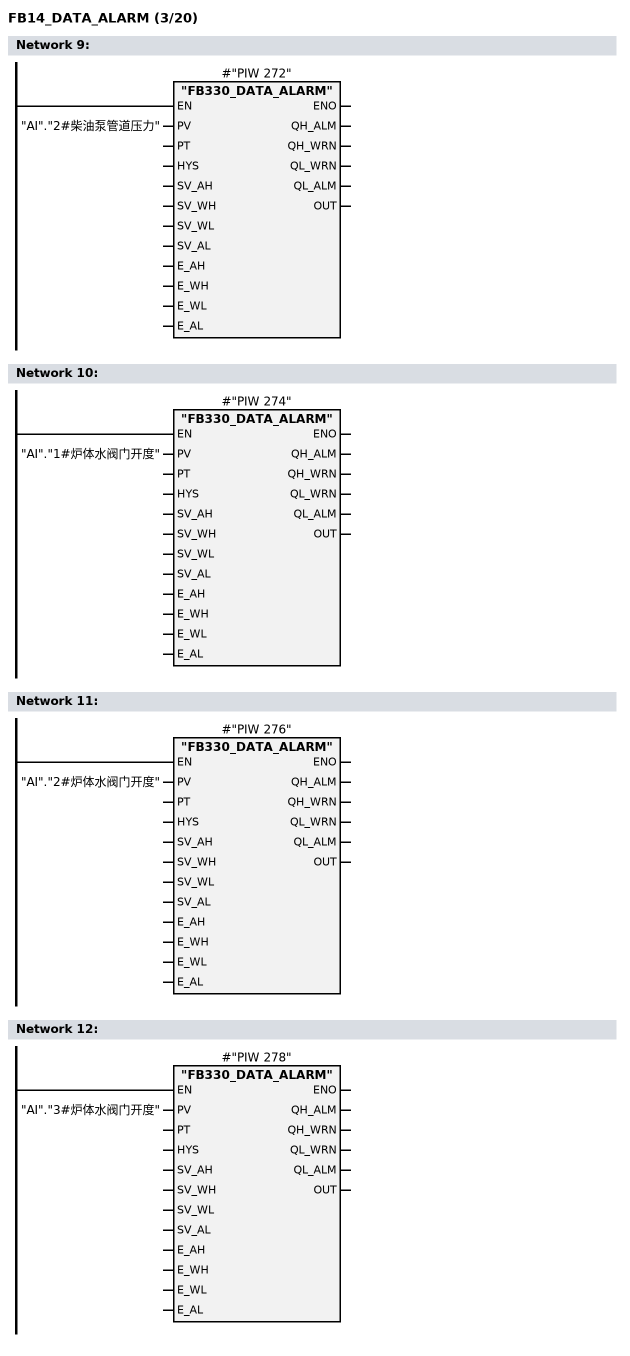
   RUNG wire#powerrail
      #"PIW 272"(PV := "AI"."2#柴油泵管道压力", PT :=, HYS :=, SV_AH :=, SV_WH :=, SV_WL :=, SV_AL :=, E_AH :=, E_WH :=, E_WL :=, E_AL :=, QH_ALM =>, QH_WRN =>, QL_WRN =>, QL_ALM =>, OUT =>)
   END_RUNG
   // the same network as SCL:
   #"PIW 272"(PV := "AI"."2#柴油泵管道压力");   // "FB330_DATA_ALARM"
END_REGION

REGION Network 10
   RUNG wire#powerrail
      #"PIW 274"(PV := "AI"."1#炉体水阀门开度", PT :=, HYS :=, SV_AH :=, SV_WH :=, SV_WL :=, SV_AL :=, E_AH :=, E_WH :=, E_WL :=, E_AL :=, QH_ALM =>, QH_WRN =>, QL_WRN =>, QL_ALM =>, OUT =>)
   END_RUNG
   // the same network as SCL:
   #"PIW 274"(PV := "AI"."1#炉体水阀门开度");   // "FB330_DATA_ALARM"
END_REGION

REGION Network 11
   RUNG wire#powerrail
      #"PIW 276"(PV := "AI"."2#炉体水阀门开度", PT :=, HYS :=, SV_AH :=, SV_WH :=, SV_WL :=, SV_AL :=, E_AH :=, E_WH :=, E_WL :=, E_AL :=, QH_ALM =>, QH_WRN =>, QL_WRN =>, QL_ALM =>, OUT =>)
   END_RUNG
   // the same network as SCL:
   #"PIW 276"(PV := "AI"."2#炉体水阀门开度");   // "FB330_DATA_ALARM"
END_REGION

REGION Network 12
   RUNG wire#powerrail
      #"PIW 278"(PV := "AI"."3#炉体水阀门开度", PT :=, HYS :=, SV_AH :=, SV_WH :=, SV_WL :=, SV_AL :=, E_AH :=, E_WH :=, E_WL :=, E_AL :=, QH_ALM =>, QH_WRN =>, QL_WRN =>, QL_ALM =>, OUT =>)
   END_RUNG
   // the same network as SCL:
   #"PIW 278"(PV := "AI"."3#炉体水阀门开度");   // "FB330_DATA_ALARM"
END_REGION

REGION Network 13
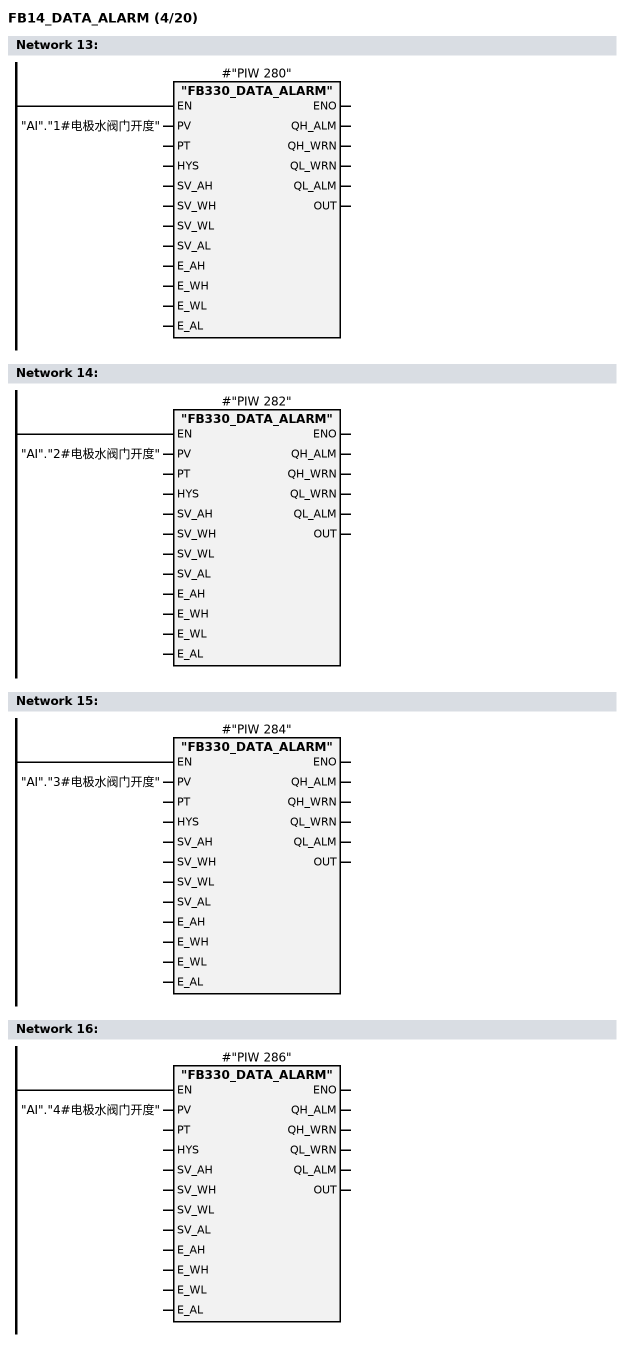
   RUNG wire#powerrail
      #"PIW 280"(PV := "AI"."1#电极水阀门开度", PT :=, HYS :=, SV_AH :=, SV_WH :=, SV_WL :=, SV_AL :=, E_AH :=, E_WH :=, E_WL :=, E_AL :=, QH_ALM =>, QH_WRN =>, QL_WRN =>, QL_ALM =>, OUT =>)
   END_RUNG
   // the same network as SCL:
   #"PIW 280"(PV := "AI"."1#电极水阀门开度");   // "FB330_DATA_ALARM"
END_REGION

REGION Network 14
   RUNG wire#powerrail
      #"PIW 282"(PV := "AI"."2#电极水阀门开度", PT :=, HYS :=, SV_AH :=, SV_WH :=, SV_WL :=, SV_AL :=, E_AH :=, E_WH :=, E_WL :=, E_AL :=, QH_ALM =>, QH_WRN =>, QL_WRN =>, QL_ALM =>, OUT =>)
   END_RUNG
   // the same network as SCL:
   #"PIW 282"(PV := "AI"."2#电极水阀门开度");   // "FB330_DATA_ALARM"
END_REGION

REGION Network 15
   RUNG wire#powerrail
      #"PIW 284"(PV := "AI"."3#电极水阀门开度", PT :=, HYS :=, SV_AH :=, SV_WH :=, SV_WL :=, SV_AL :=, E_AH :=, E_WH :=, E_WL :=, E_AL :=, QH_ALM =>, QH_WRN =>, QL_WRN =>, QL_ALM =>, OUT =>)
   END_RUNG
   // the same network as SCL:
   #"PIW 284"(PV := "AI"."3#电极水阀门开度");   // "FB330_DATA_ALARM"
END_REGION

REGION Network 16
   RUNG wire#powerrail
      #"PIW 286"(PV := "AI"."4#电极水阀门开度", PT :=, HYS :=, SV_AH :=, SV_WH :=, SV_WL :=, SV_AL :=, E_AH :=, E_WH :=, E_WL :=, E_AL :=, QH_ALM =>, QH_WRN =>, QL_WRN =>, QL_ALM =>, OUT =>)
   END_RUNG
   // the same network as SCL:
   #"PIW 286"(PV := "AI"."4#电极水阀门开度");   // "FB330_DATA_ALARM"
END_REGION

REGION Network 17
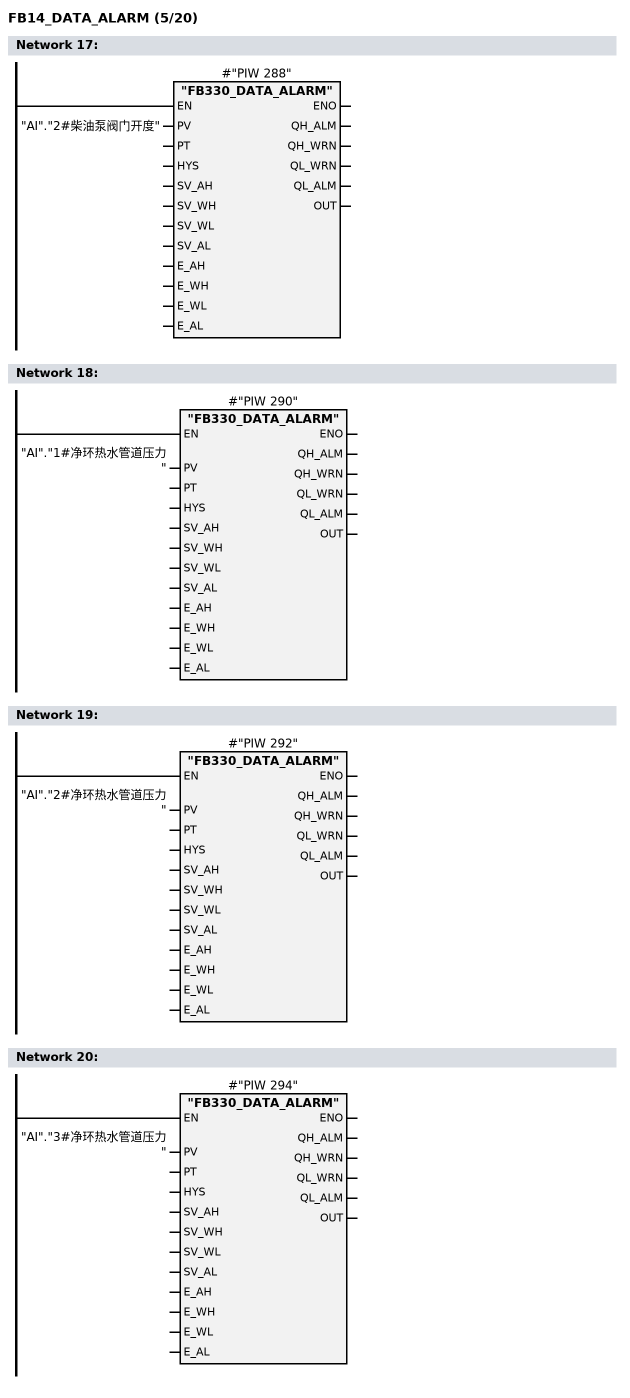
   RUNG wire#powerrail
      #"PIW 288"(PV := "AI"."2#柴油泵阀门开度", PT :=, HYS :=, SV_AH :=, SV_WH :=, SV_WL :=, SV_AL :=, E_AH :=, E_WH :=, E_WL :=, E_AL :=, QH_ALM =>, QH_WRN =>, QL_WRN =>, QL_ALM =>, OUT =>)
   END_RUNG
   // the same network as SCL:
   #"PIW 288"(PV := "AI"."2#柴油泵阀门开度");   // "FB330_DATA_ALARM"
END_REGION

REGION Network 18
   RUNG wire#powerrail
      #"PIW 290"(PV := "AI"."1#净环热水管道压力", PT :=, HYS :=, SV_AH :=, SV_WH :=, SV_WL :=, SV_AL :=, E_AH :=, E_WH :=, E_WL :=, E_AL :=, QH_ALM =>, QH_WRN =>, QL_WRN =>, QL_ALM =>, OUT =>)
   END_RUNG
   // the same network as SCL:
   #"PIW 290"(PV := "AI"."1#净环热水管道压力");   // "FB330_DATA_ALARM"
END_REGION

REGION Network 19
   RUNG wire#powerrail
      #"PIW 292"(PV := "AI"."2#净环热水管道压力", PT :=, HYS :=, SV_AH :=, SV_WH :=, SV_WL :=, SV_AL :=, E_AH :=, E_WH :=, E_WL :=, E_AL :=, QH_ALM =>, QH_WRN =>, QL_WRN =>, QL_ALM =>, OUT =>)
   END_RUNG
   // the same network as SCL:
   #"PIW 292"(PV := "AI"."2#净环热水管道压力");   // "FB330_DATA_ALARM"
END_REGION

REGION Network 20
   RUNG wire#powerrail
      #"PIW 294"(PV := "AI"."3#净环热水管道压力", PT :=, HYS :=, SV_AH :=, SV_WH :=, SV_WL :=, SV_AL :=, E_AH :=, E_WH :=, E_WL :=, E_AL :=, QH_ALM =>, QH_WRN =>, QL_WRN =>, QL_ALM =>, OUT =>)
   END_RUNG
   // the same network as SCL:
   #"PIW 294"(PV := "AI"."3#净环热水管道压力");   // "FB330_DATA_ALARM"
END_REGION

REGION Network 21
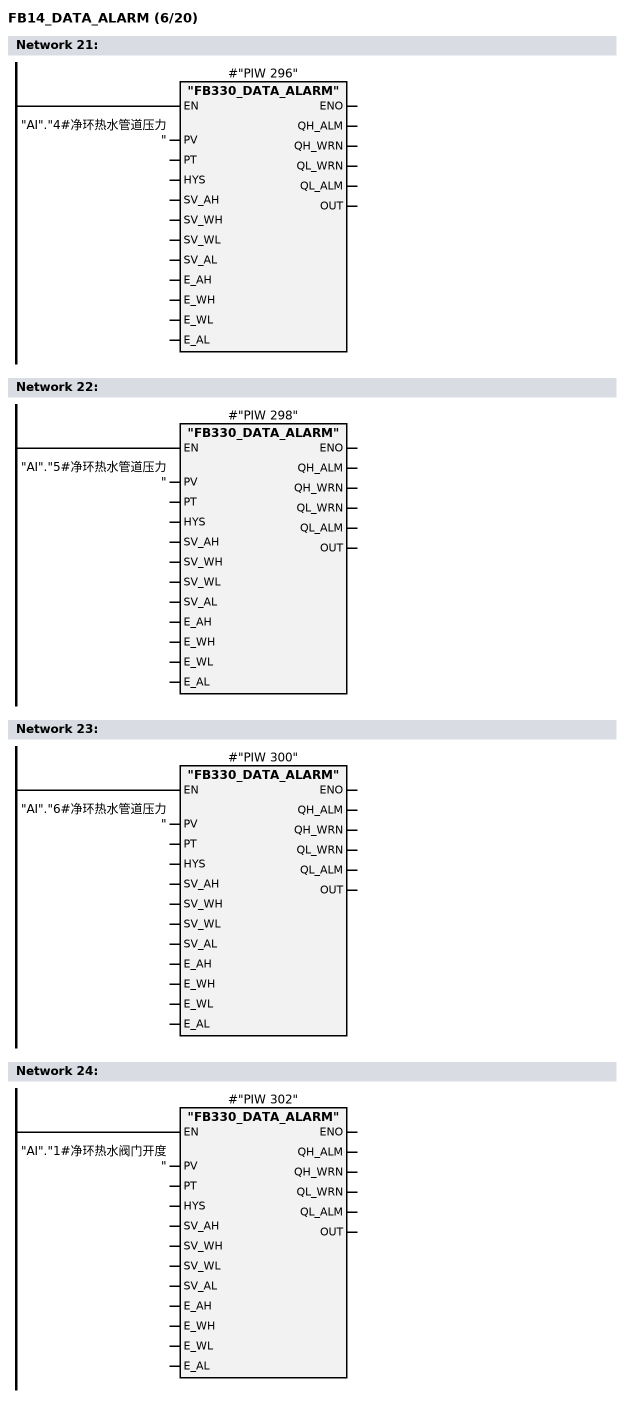
   RUNG wire#powerrail
      #"PIW 296"(PV := "AI"."4#净环热水管道压力", PT :=, HYS :=, SV_AH :=, SV_WH :=, SV_WL :=, SV_AL :=, E_AH :=, E_WH :=, E_WL :=, E_AL :=, QH_ALM =>, QH_WRN =>, QL_WRN =>, QL_ALM =>, OUT =>)
   END_RUNG
   // the same network as SCL:
   #"PIW 296"(PV := "AI"."4#净环热水管道压力");   // "FB330_DATA_ALARM"
END_REGION

REGION Network 22
   RUNG wire#powerrail
      #"PIW 298"(PV := "AI"."5#净环热水管道压力", PT :=, HYS :=, SV_AH :=, SV_WH :=, SV_WL :=, SV_AL :=, E_AH :=, E_WH :=, E_WL :=, E_AL :=, QH_ALM =>, QH_WRN =>, QL_WRN =>, QL_ALM =>, OUT =>)
   END_RUNG
   // the same network as SCL:
   #"PIW 298"(PV := "AI"."5#净环热水管道压力");   // "FB330_DATA_ALARM"
END_REGION

REGION Network 23
   RUNG wire#powerrail
      #"PIW 300"(PV := "AI"."6#净环热水管道压力", PT :=, HYS :=, SV_AH :=, SV_WH :=, SV_WL :=, SV_AL :=, E_AH :=, E_WH :=, E_WL :=, E_AL :=, QH_ALM =>, QH_WRN =>, QL_WRN =>, QL_ALM =>, OUT =>)
   END_RUNG
   // the same network as SCL:
   #"PIW 300"(PV := "AI"."6#净环热水管道压力");   // "FB330_DATA_ALARM"
END_REGION

REGION Network 24
   RUNG wire#powerrail
      #"PIW 302"(PV := "AI"."1#净环热水阀门开度", PT :=, HYS :=, SV_AH :=, SV_WH :=, SV_WL :=, SV_AL :=, E_AH :=, E_WH :=, E_WL :=, E_AL :=, QH_ALM =>, QH_WRN =>, QL_WRN =>, QL_ALM =>, OUT =>)
   END_RUNG
   // the same network as SCL:
   #"PIW 302"(PV := "AI"."1#净环热水阀门开度");   // "FB330_DATA_ALARM"
END_REGION

REGION Network 25
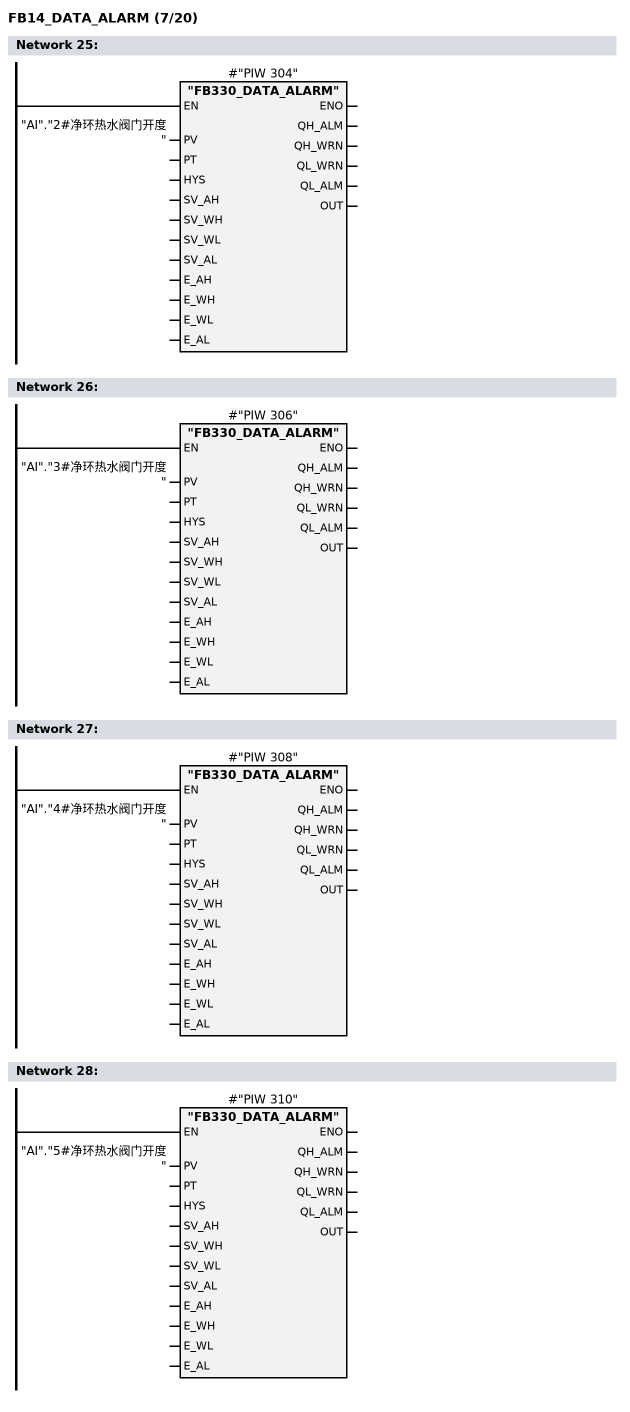
   RUNG wire#powerrail
      #"PIW 304"(PV := "AI"."2#净环热水阀门开度", PT :=, HYS :=, SV_AH :=, SV_WH :=, SV_WL :=, SV_AL :=, E_AH :=, E_WH :=, E_WL :=, E_AL :=, QH_ALM =>, QH_WRN =>, QL_WRN =>, QL_ALM =>, OUT =>)
   END_RUNG
   // the same network as SCL:
   #"PIW 304"(PV := "AI"."2#净环热水阀门开度");   // "FB330_DATA_ALARM"
END_REGION

REGION Network 26
   RUNG wire#powerrail
      #"PIW 306"(PV := "AI"."3#净环热水阀门开度", PT :=, HYS :=, SV_AH :=, SV_WH :=, SV_WL :=, SV_AL :=, E_AH :=, E_WH :=, E_WL :=, E_AL :=, QH_ALM =>, QH_WRN =>, QL_WRN =>, QL_ALM =>, OUT =>)
   END_RUNG
   // the same network as SCL:
   #"PIW 306"(PV := "AI"."3#净环热水阀门开度");   // "FB330_DATA_ALARM"
END_REGION

REGION Network 27
   RUNG wire#powerrail
      #"PIW 308"(PV := "AI"."4#净环热水阀门开度", PT :=, HYS :=, SV_AH :=, SV_WH :=, SV_WL :=, SV_AL :=, E_AH :=, E_WH :=, E_WL :=, E_AL :=, QH_ALM =>, QH_WRN =>, QL_WRN =>, QL_ALM =>, OUT =>)
   END_RUNG
   // the same network as SCL:
   #"PIW 308"(PV := "AI"."4#净环热水阀门开度");   // "FB330_DATA_ALARM"
END_REGION

REGION Network 28
   RUNG wire#powerrail
      #"PIW 310"(PV := "AI"."5#净环热水阀门开度", PT :=, HYS :=, SV_AH :=, SV_WH :=, SV_WL :=, SV_AL :=, E_AH :=, E_WH :=, E_WL :=, E_AL :=, QH_ALM =>, QH_WRN =>, QL_WRN =>, QL_ALM =>, OUT =>)
   END_RUNG
   // the same network as SCL:
   #"PIW 310"(PV := "AI"."5#净环热水阀门开度");   // "FB330_DATA_ALARM"
END_REGION

REGION Network 29
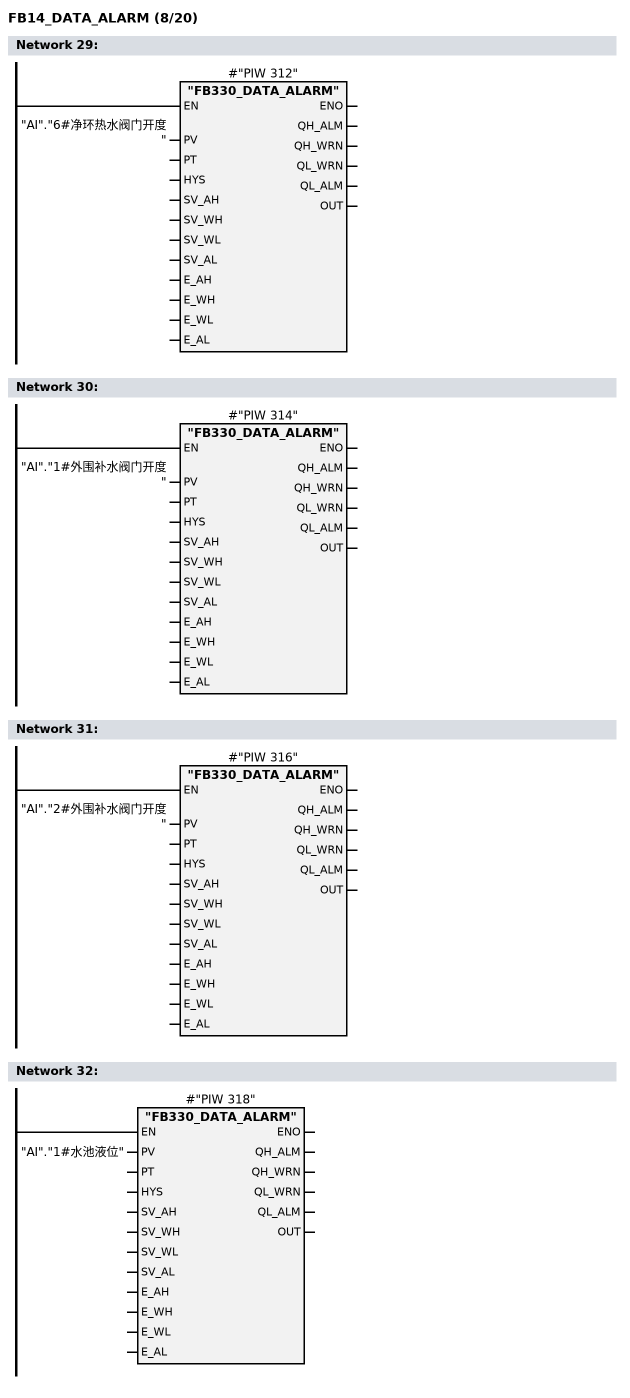
   RUNG wire#powerrail
      #"PIW 312"(PV := "AI"."6#净环热水阀门开度", PT :=, HYS :=, SV_AH :=, SV_WH :=, SV_WL :=, SV_AL :=, E_AH :=, E_WH :=, E_WL :=, E_AL :=, QH_ALM =>, QH_WRN =>, QL_WRN =>, QL_ALM =>, OUT =>)
   END_RUNG
   // the same network as SCL:
   #"PIW 312"(PV := "AI"."6#净环热水阀门开度");   // "FB330_DATA_ALARM"
END_REGION

REGION Network 30
   RUNG wire#powerrail
      #"PIW 314"(PV := "AI"."1#外围补水阀门开度", PT :=, HYS :=, SV_AH :=, SV_WH :=, SV_WL :=, SV_AL :=, E_AH :=, E_WH :=, E_WL :=, E_AL :=, QH_ALM =>, QH_WRN =>, QL_WRN =>, QL_ALM =>, OUT =>)
   END_RUNG
   // the same network as SCL:
   #"PIW 314"(PV := "AI"."1#外围补水阀门开度");   // "FB330_DATA_ALARM"
END_REGION

REGION Network 31
   RUNG wire#powerrail
      #"PIW 316"(PV := "AI"."2#外围补水阀门开度", PT :=, HYS :=, SV_AH :=, SV_WH :=, SV_WL :=, SV_AL :=, E_AH :=, E_WH :=, E_WL :=, E_AL :=, QH_ALM =>, QH_WRN =>, QL_WRN =>, QL_ALM =>, OUT =>)
   END_RUNG
   // the same network as SCL:
   #"PIW 316"(PV := "AI"."2#外围补水阀门开度");   // "FB330_DATA_ALARM"
END_REGION

REGION Network 32
   RUNG wire#powerrail
      #"PIW 318"(PV := "AI"."1#水池液位", PT :=, HYS :=, SV_AH :=, SV_WH :=, SV_WL :=, SV_AL :=, E_AH :=, E_WH :=, E_WL :=, E_AL :=, QH_ALM =>, QH_WRN =>, QL_WRN =>, QL_ALM =>, OUT =>)
   END_RUNG
   // the same network as SCL:
   #"PIW 318"(PV := "AI"."1#水池液位");   // "FB330_DATA_ALARM"
END_REGION

REGION Network 33
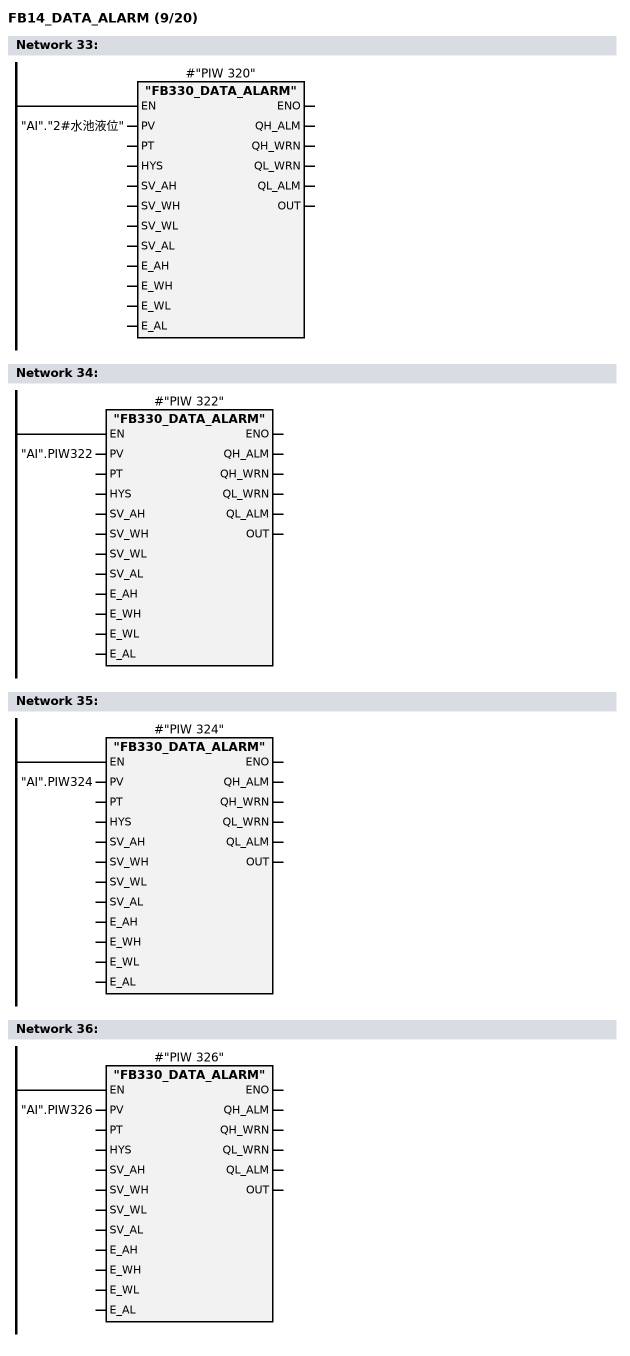
   RUNG wire#powerrail
      #"PIW 320"(PV := "AI"."2#水池液位", PT :=, HYS :=, SV_AH :=, SV_WH :=, SV_WL :=, SV_AL :=, E_AH :=, E_WH :=, E_WL :=, E_AL :=, QH_ALM =>, QH_WRN =>, QL_WRN =>, QL_ALM =>, OUT =>)
   END_RUNG
   // the same network as SCL:
   #"PIW 320"(PV := "AI"."2#水池液位");   // "FB330_DATA_ALARM"
END_REGION

REGION Network 34
   RUNG wire#powerrail
      #"PIW 322"(PV := "AI".PIW322, PT :=, HYS :=, SV_AH :=, SV_WH :=, SV_WL :=, SV_AL :=, E_AH :=, E_WH :=, E_WL :=, E_AL :=, QH_ALM =>, QH_WRN =>, QL_WRN =>, QL_ALM =>, OUT =>)
   END_RUNG
   // the same network as SCL:
   #"PIW 322"(PV := "AI".PIW322);   // "FB330_DATA_ALARM"
END_REGION

REGION Network 35
   RUNG wire#powerrail
      #"PIW 324"(PV := "AI".PIW324, PT :=, HYS :=, SV_AH :=, SV_WH :=, SV_WL :=, SV_AL :=, E_AH :=, E_WH :=, E_WL :=, E_AL :=, QH_ALM =>, QH_WRN =>, QL_WRN =>, QL_ALM =>, OUT =>)
   END_RUNG
   // the same network as SCL:
   #"PIW 324"(PV := "AI".PIW324);   // "FB330_DATA_ALARM"
END_REGION

REGION Network 36
   RUNG wire#powerrail
      #"PIW 326"(PV := "AI".PIW326, PT :=, HYS :=, SV_AH :=, SV_WH :=, SV_WL :=, SV_AL :=, E_AH :=, E_WH :=, E_WL :=, E_AL :=, QH_ALM =>, QH_WRN =>, QL_WRN =>, QL_ALM =>, OUT =>)
   END_RUNG
   // the same network as SCL:
   #"PIW 326"(PV := "AI".PIW326);   // "FB330_DATA_ALARM"
END_REGION

REGION Network 37
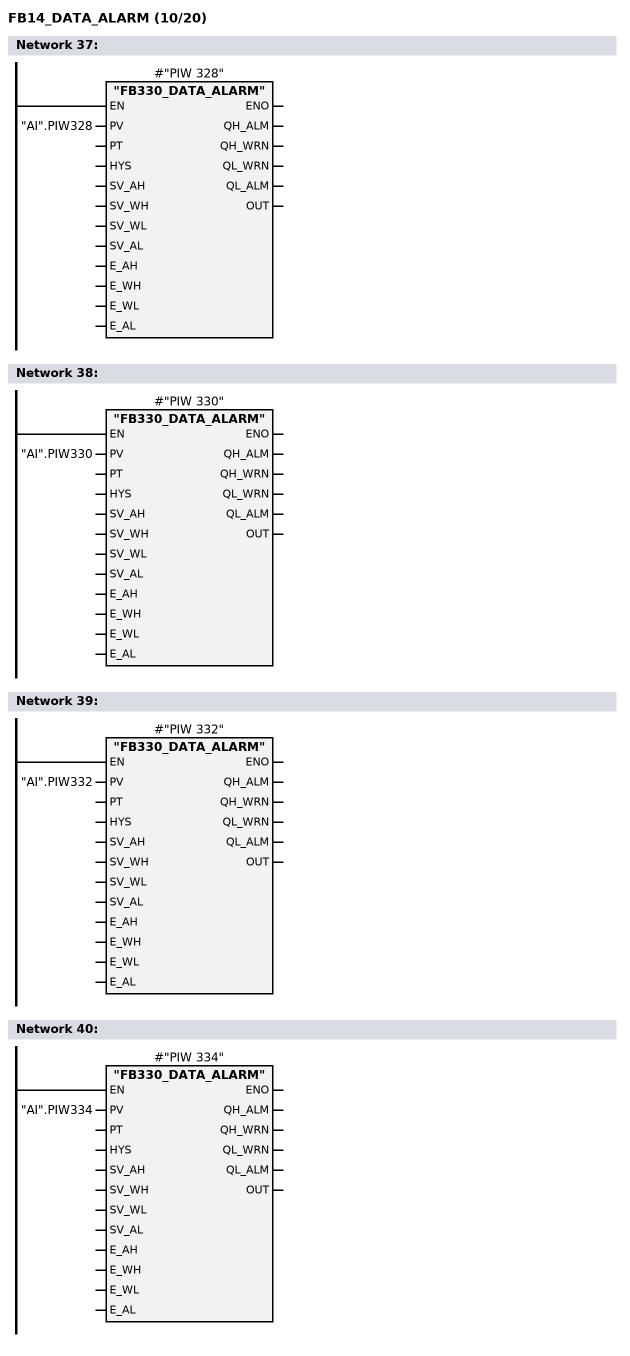
   RUNG wire#powerrail
      #"PIW 328"(PV := "AI".PIW328, PT :=, HYS :=, SV_AH :=, SV_WH :=, SV_WL :=, SV_AL :=, E_AH :=, E_WH :=, E_WL :=, E_AL :=, QH_ALM =>, QH_WRN =>, QL_WRN =>, QL_ALM =>, OUT =>)
   END_RUNG
   // the same network as SCL:
   #"PIW 328"(PV := "AI".PIW328);   // "FB330_DATA_ALARM"
END_REGION

REGION Network 38
   RUNG wire#powerrail
      #"PIW 330"(PV := "AI".PIW330, PT :=, HYS :=, SV_AH :=, SV_WH :=, SV_WL :=, SV_AL :=, E_AH :=, E_WH :=, E_WL :=, E_AL :=, QH_ALM =>, QH_WRN =>, QL_WRN =>, QL_ALM =>, OUT =>)
   END_RUNG
   // the same network as SCL:
   #"PIW 330"(PV := "AI".PIW330);   // "FB330_DATA_ALARM"
END_REGION

REGION Network 39
   RUNG wire#powerrail
      #"PIW 332"(PV := "AI".PIW332, PT :=, HYS :=, SV_AH :=, SV_WH :=, SV_WL :=, SV_AL :=, E_AH :=, E_WH :=, E_WL :=, E_AL :=, QH_ALM =>, QH_WRN =>, QL_WRN =>, QL_ALM =>, OUT =>)
   END_RUNG
   // the same network as SCL:
   #"PIW 332"(PV := "AI".PIW332);   // "FB330_DATA_ALARM"
END_REGION

REGION Network 40
   RUNG wire#powerrail
      #"PIW 334"(PV := "AI".PIW334, PT :=, HYS :=, SV_AH :=, SV_WH :=, SV_WL :=, SV_AL :=, E_AH :=, E_WH :=, E_WL :=, E_AL :=, QH_ALM =>, QH_WRN =>, QL_WRN =>, QL_ALM =>, OUT =>)
   END_RUNG
   // the same network as SCL:
   #"PIW 334"(PV := "AI".PIW334);   // "FB330_DATA_ALARM"
END_REGION

REGION Network 41
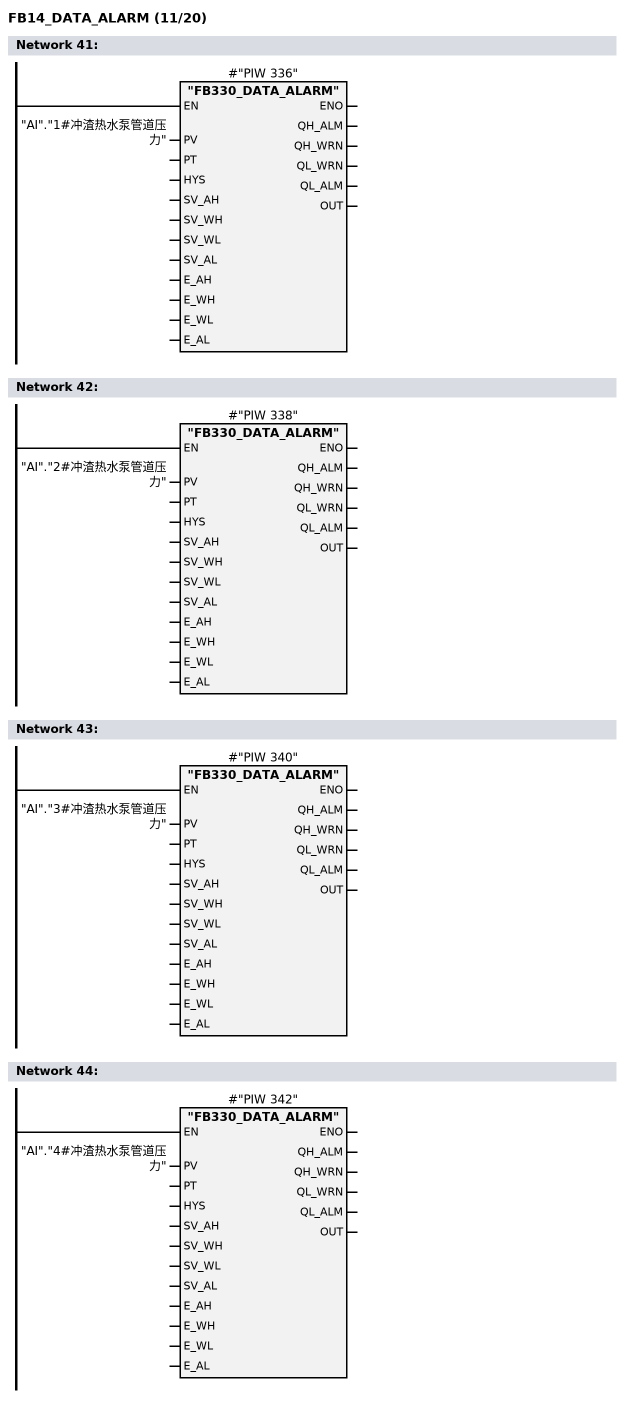
   RUNG wire#powerrail
      #"PIW 336"(PV := "AI"."1#冲渣热水泵管道压力", PT :=, HYS :=, SV_AH :=, SV_WH :=, SV_WL :=, SV_AL :=, E_AH :=, E_WH :=, E_WL :=, E_AL :=, QH_ALM =>, QH_WRN =>, QL_WRN =>, QL_ALM =>, OUT =>)
   END_RUNG
   // the same network as SCL:
   #"PIW 336"(PV := "AI"."1#冲渣热水泵管道压力");   // "FB330_DATA_ALARM"
END_REGION

REGION Network 42
   RUNG wire#powerrail
      #"PIW 338"(PV := "AI"."2#冲渣热水泵管道压力", PT :=, HYS :=, SV_AH :=, SV_WH :=, SV_WL :=, SV_AL :=, E_AH :=, E_WH :=, E_WL :=, E_AL :=, QH_ALM =>, QH_WRN =>, QL_WRN =>, QL_ALM =>, OUT =>)
   END_RUNG
   // the same network as SCL:
   #"PIW 338"(PV := "AI"."2#冲渣热水泵管道压力");   // "FB330_DATA_ALARM"
END_REGION

REGION Network 43
   RUNG wire#powerrail
      #"PIW 340"(PV := "AI"."3#冲渣热水泵管道压力", PT :=, HYS :=, SV_AH :=, SV_WH :=, SV_WL :=, SV_AL :=, E_AH :=, E_WH :=, E_WL :=, E_AL :=, QH_ALM =>, QH_WRN =>, QL_WRN =>, QL_ALM =>, OUT =>)
   END_RUNG
   // the same network as SCL:
   #"PIW 340"(PV := "AI"."3#冲渣热水泵管道压力");   // "FB330_DATA_ALARM"
END_REGION

REGION Network 44
   RUNG wire#powerrail
      #"PIW 342"(PV := "AI"."4#冲渣热水泵管道压力", PT :=, HYS :=, SV_AH :=, SV_WH :=, SV_WL :=, SV_AL :=, E_AH :=, E_WH :=, E_WL :=, E_AL :=, QH_ALM =>, QH_WRN =>, QL_WRN =>, QL_ALM =>, OUT =>)
   END_RUNG
   // the same network as SCL:
   #"PIW 342"(PV := "AI"."4#冲渣热水泵管道压力");   // "FB330_DATA_ALARM"
END_REGION

REGION Network 45
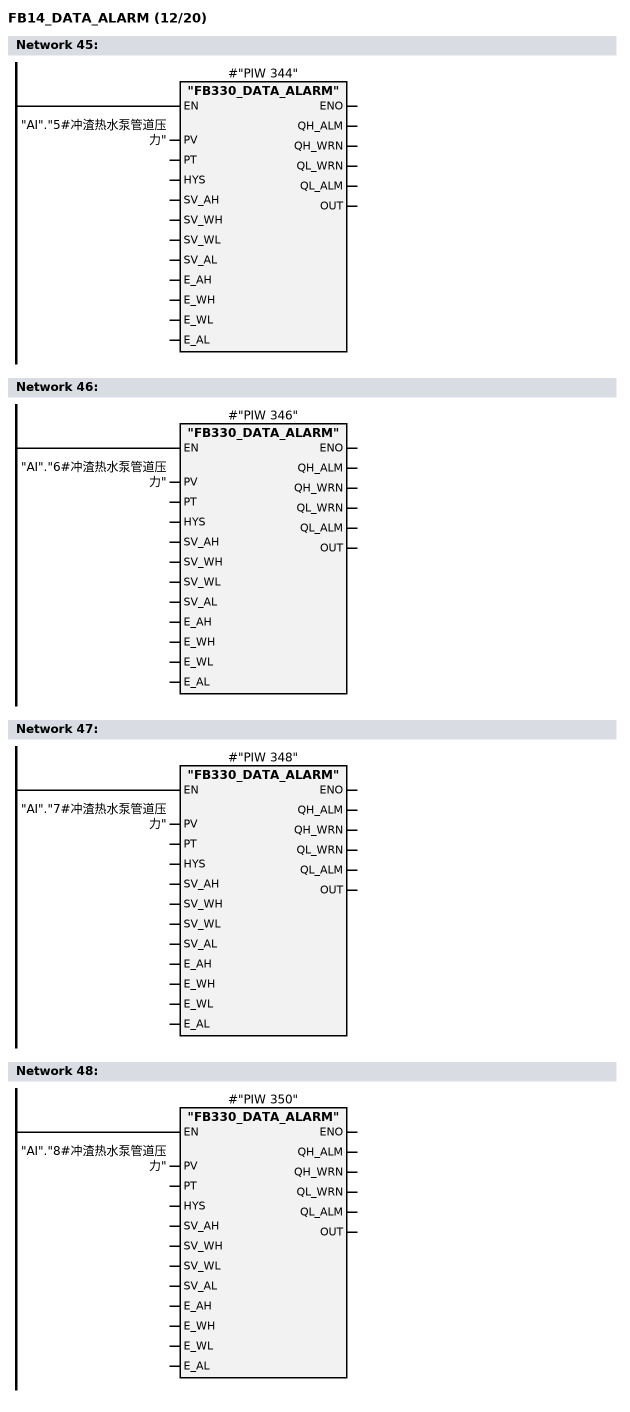
   RUNG wire#powerrail
      #"PIW 344"(PV := "AI"."5#冲渣热水泵管道压力", PT :=, HYS :=, SV_AH :=, SV_WH :=, SV_WL :=, SV_AL :=, E_AH :=, E_WH :=, E_WL :=, E_AL :=, QH_ALM =>, QH_WRN =>, QL_WRN =>, QL_ALM =>, OUT =>)
   END_RUNG
   // the same network as SCL:
   #"PIW 344"(PV := "AI"."5#冲渣热水泵管道压力");   // "FB330_DATA_ALARM"
END_REGION

REGION Network 46
   RUNG wire#powerrail
      #"PIW 346"(PV := "AI"."6#冲渣热水泵管道压力", PT :=, HYS :=, SV_AH :=, SV_WH :=, SV_WL :=, SV_AL :=, E_AH :=, E_WH :=, E_WL :=, E_AL :=, QH_ALM =>, QH_WRN =>, QL_WRN =>, QL_ALM =>, OUT =>)
   END_RUNG
   // the same network as SCL:
   #"PIW 346"(PV := "AI"."6#冲渣热水泵管道压力");   // "FB330_DATA_ALARM"
END_REGION

REGION Network 47
   RUNG wire#powerrail
      #"PIW 348"(PV := "AI"."7#冲渣热水泵管道压力", PT :=, HYS :=, SV_AH :=, SV_WH :=, SV_WL :=, SV_AL :=, E_AH :=, E_WH :=, E_WL :=, E_AL :=, QH_ALM =>, QH_WRN =>, QL_WRN =>, QL_ALM =>, OUT =>)
   END_RUNG
   // the same network as SCL:
   #"PIW 348"(PV := "AI"."7#冲渣热水泵管道压力");   // "FB330_DATA_ALARM"
END_REGION

REGION Network 48
   RUNG wire#powerrail
      #"PIW 350"(PV := "AI"."8#冲渣热水泵管道压力", PT :=, HYS :=, SV_AH :=, SV_WH :=, SV_WL :=, SV_AL :=, E_AH :=, E_WH :=, E_WL :=, E_AL :=, QH_ALM =>, QH_WRN =>, QL_WRN =>, QL_ALM =>, OUT =>)
   END_RUNG
   // the same network as SCL:
   #"PIW 350"(PV := "AI"."8#冲渣热水泵管道压力");   // "FB330_DATA_ALARM"
END_REGION

REGION Network 49
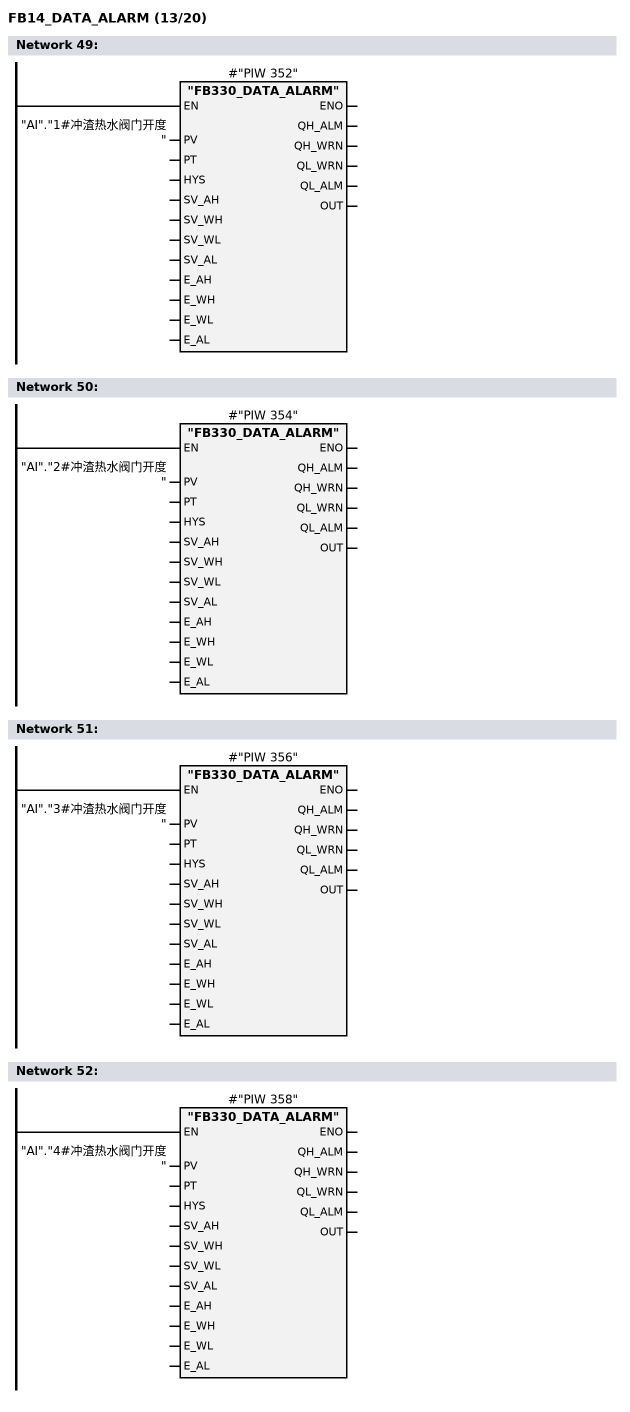
   RUNG wire#powerrail
      #"PIW 352"(PV := "AI"."1#冲渣热水阀门开度", PT :=, HYS :=, SV_AH :=, SV_WH :=, SV_WL :=, SV_AL :=, E_AH :=, E_WH :=, E_WL :=, E_AL :=, QH_ALM =>, QH_WRN =>, QL_WRN =>, QL_ALM =>, OUT =>)
   END_RUNG
   // the same network as SCL:
   #"PIW 352"(PV := "AI"."1#冲渣热水阀门开度");   // "FB330_DATA_ALARM"
END_REGION

REGION Network 50
   RUNG wire#powerrail
      #"PIW 354"(PV := "AI"."2#冲渣热水阀门开度", PT :=, HYS :=, SV_AH :=, SV_WH :=, SV_WL :=, SV_AL :=, E_AH :=, E_WH :=, E_WL :=, E_AL :=, QH_ALM =>, QH_WRN =>, QL_WRN =>, QL_ALM =>, OUT =>)
   END_RUNG
   // the same network as SCL:
   #"PIW 354"(PV := "AI"."2#冲渣热水阀门开度");   // "FB330_DATA_ALARM"
END_REGION

REGION Network 51
   RUNG wire#powerrail
      #"PIW 356"(PV := "AI"."3#冲渣热水阀门开度", PT :=, HYS :=, SV_AH :=, SV_WH :=, SV_WL :=, SV_AL :=, E_AH :=, E_WH :=, E_WL :=, E_AL :=, QH_ALM =>, QH_WRN =>, QL_WRN =>, QL_ALM =>, OUT =>)
   END_RUNG
   // the same network as SCL:
   #"PIW 356"(PV := "AI"."3#冲渣热水阀门开度");   // "FB330_DATA_ALARM"
END_REGION

REGION Network 52
   RUNG wire#powerrail
      #"PIW 358"(PV := "AI"."4#冲渣热水阀门开度", PT :=, HYS :=, SV_AH :=, SV_WH :=, SV_WL :=, SV_AL :=, E_AH :=, E_WH :=, E_WL :=, E_AL :=, QH_ALM =>, QH_WRN =>, QL_WRN =>, QL_ALM =>, OUT =>)
   END_RUNG
   // the same network as SCL:
   #"PIW 358"(PV := "AI"."4#冲渣热水阀门开度");   // "FB330_DATA_ALARM"
END_REGION

REGION Network 53
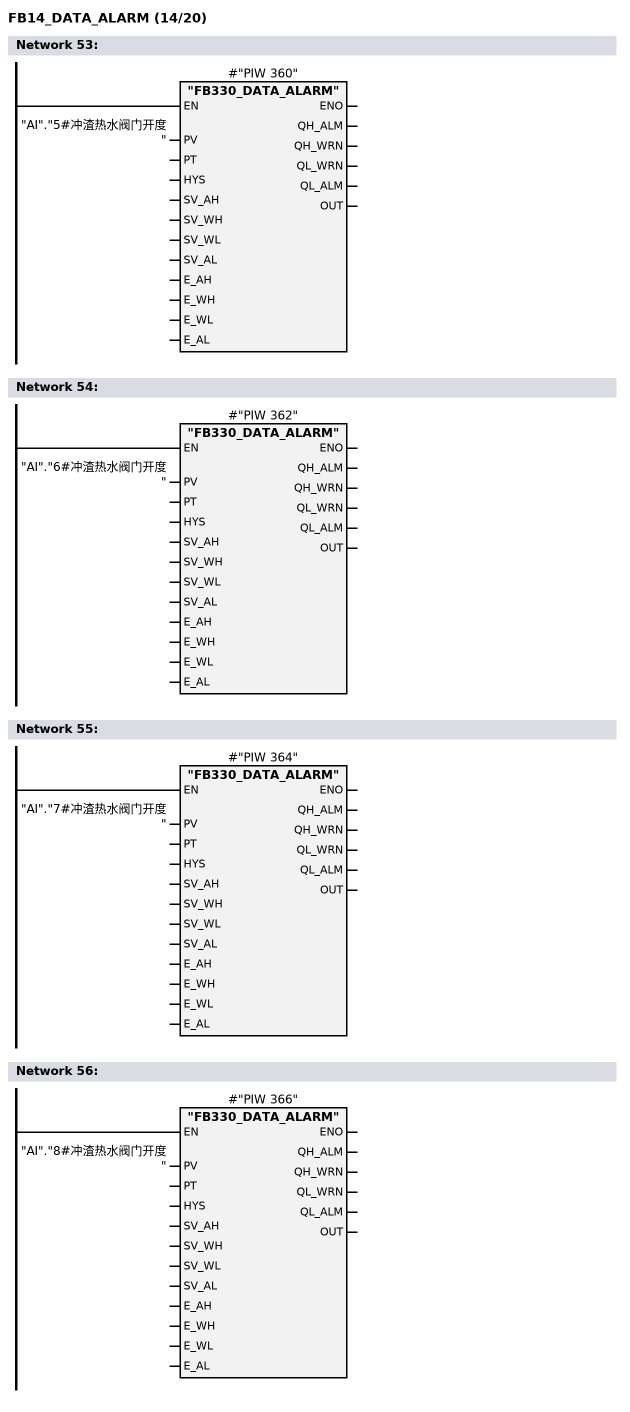
   RUNG wire#powerrail
      #"PIW 360"(PV := "AI"."5#冲渣热水阀门开度", PT :=, HYS :=, SV_AH :=, SV_WH :=, SV_WL :=, SV_AL :=, E_AH :=, E_WH :=, E_WL :=, E_AL :=, QH_ALM =>, QH_WRN =>, QL_WRN =>, QL_ALM =>, OUT =>)
   END_RUNG
   // the same network as SCL:
   #"PIW 360"(PV := "AI"."5#冲渣热水阀门开度");   // "FB330_DATA_ALARM"
END_REGION

REGION Network 54
   RUNG wire#powerrail
      #"PIW 362"(PV := "AI"."6#冲渣热水阀门开度", PT :=, HYS :=, SV_AH :=, SV_WH :=, SV_WL :=, SV_AL :=, E_AH :=, E_WH :=, E_WL :=, E_AL :=, QH_ALM =>, QH_WRN =>, QL_WRN =>, QL_ALM =>, OUT =>)
   END_RUNG
   // the same network as SCL:
   #"PIW 362"(PV := "AI"."6#冲渣热水阀门开度");   // "FB330_DATA_ALARM"
END_REGION

REGION Network 55
   RUNG wire#powerrail
      #"PIW 364"(PV := "AI"."7#冲渣热水阀门开度", PT :=, HYS :=, SV_AH :=, SV_WH :=, SV_WL :=, SV_AL :=, E_AH :=, E_WH :=, E_WL :=, E_AL :=, QH_ALM =>, QH_WRN =>, QL_WRN =>, QL_ALM =>, OUT =>)
   END_RUNG
   // the same network as SCL:
   #"PIW 364"(PV := "AI"."7#冲渣热水阀门开度");   // "FB330_DATA_ALARM"
END_REGION

REGION Network 56
   RUNG wire#powerrail
      #"PIW 366"(PV := "AI"."8#冲渣热水阀门开度", PT :=, HYS :=, SV_AH :=, SV_WH :=, SV_WL :=, SV_AL :=, E_AH :=, E_WH :=, E_WL :=, E_AL :=, QH_ALM =>, QH_WRN =>, QL_WRN =>, QL_ALM =>, OUT =>)
   END_RUNG
   // the same network as SCL:
   #"PIW 366"(PV := "AI"."8#冲渣热水阀门开度");   // "FB330_DATA_ALARM"
END_REGION

REGION Network 57
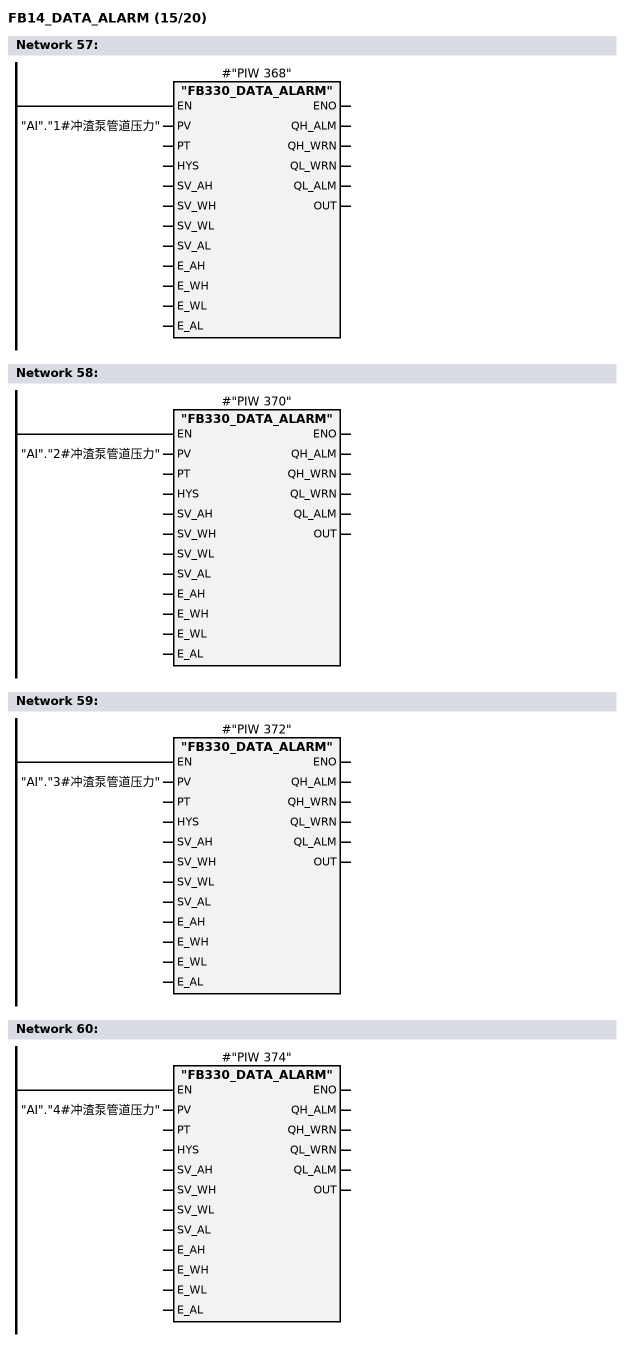
   RUNG wire#powerrail
      #"PIW 368"(PV := "AI"."1#冲渣泵管道压力", PT :=, HYS :=, SV_AH :=, SV_WH :=, SV_WL :=, SV_AL :=, E_AH :=, E_WH :=, E_WL :=, E_AL :=, QH_ALM =>, QH_WRN =>, QL_WRN =>, QL_ALM =>, OUT =>)
   END_RUNG
   // the same network as SCL:
   #"PIW 368"(PV := "AI"."1#冲渣泵管道压力");   // "FB330_DATA_ALARM"
END_REGION

REGION Network 58
   RUNG wire#powerrail
      #"PIW 370"(PV := "AI"."2#冲渣泵管道压力", PT :=, HYS :=, SV_AH :=, SV_WH :=, SV_WL :=, SV_AL :=, E_AH :=, E_WH :=, E_WL :=, E_AL :=, QH_ALM =>, QH_WRN =>, QL_WRN =>, QL_ALM =>, OUT =>)
   END_RUNG
   // the same network as SCL:
   #"PIW 370"(PV := "AI"."2#冲渣泵管道压力");   // "FB330_DATA_ALARM"
END_REGION

REGION Network 59
   RUNG wire#powerrail
      #"PIW 372"(PV := "AI"."3#冲渣泵管道压力", PT :=, HYS :=, SV_AH :=, SV_WH :=, SV_WL :=, SV_AL :=, E_AH :=, E_WH :=, E_WL :=, E_AL :=, QH_ALM =>, QH_WRN =>, QL_WRN =>, QL_ALM =>, OUT =>)
   END_RUNG
   // the same network as SCL:
   #"PIW 372"(PV := "AI"."3#冲渣泵管道压力");   // "FB330_DATA_ALARM"
END_REGION

REGION Network 60
   RUNG wire#powerrail
      #"PIW 374"(PV := "AI"."4#冲渣泵管道压力", PT :=, HYS :=, SV_AH :=, SV_WH :=, SV_WL :=, SV_AL :=, E_AH :=, E_WH :=, E_WL :=, E_AL :=, QH_ALM =>, QH_WRN =>, QL_WRN =>, QL_ALM =>, OUT =>)
   END_RUNG
   // the same network as SCL:
   #"PIW 374"(PV := "AI"."4#冲渣泵管道压力");   // "FB330_DATA_ALARM"
END_REGION

REGION Network 61
